IF NOT m_xInitial THEN
	BarCylinderIO.tLoadDelay:=T#3s;
	m_xInitial:=1;
END_IF;
IF g_xManual THEN    (*手动*)
	BarCylinderIO.xNextRun:=0;
	BarCylinderIO.xBarCylinder:=BarCylinderIO.xBarCylinderButton;
	BarCylinderIO.xBarCylinderSecondary	:=BarCylinderIO.xBarSecondaryButton;
	BarCylinderIO.xTransportMotorCW:= BarCylinderIO.xTransportMotorCWButton 
																	AND NOT BarCylinderIO.xTransportMotorCCWButton 
																	AND NOT BarCylinderIO.xTransportMotorCCW ;
	BarCylinderIO.xTransportMotorCCW:=BarCylinderIO.xTransportMotorCCWButton 
																		AND NOT BarCylinderIO.xTransportMotorCWButton 
																		AND NOT BarCylinderIO.xTransportMotorCW;
END_IF;
IF g_xAuto THEN(*自动*)
    IF BarCylinderIO.xUnload   (*下料*)
    	AND NOT BarCylinderIO.xEmpty  (*有料*)
    	AND NOT BarCylinderIO.xNextRun  (*下段线体旋转*)
    	AND NOT (g_xResetSingle AND BarCylinderIO.iDeviceID=g_iDeviceIDSelect)(*无复位信号*)
    	THEN(*收到卸料命令，当阻挡器不为空时*)
    	BarCylinderIO.xBarCylinder:=1;
    	BarCylinderIO.xNextRun:=1;(*确保下料命令只执行一次，防止物料在输送过程中又有卸料命令导致多次卸料*)
    	BarCylinderIO.xTransportMotorCW:=1;
    END_IF;
    IF NOT  BarCylinderIO.xUnload  THEN
    	BarCylinderIO.xNextRun:=0;
    	BarCylinderIO.xBarCylinder:=0;
    END_IF;
    m_tonLoadDelay(IN:= BarCylinderIO.xPresentSwitch ,PT:= BarCylinderIO.tLoadDelay ,Q:= m_xLoadDelay,ET:= m_tLoadDelayCurrentTime );
    IF m_xLoadDelay OR  BarCylinderIO.xNextRun  THEN
    	BarCylinderIO.xEmpty:=0;
    	BarCylinderIO.xBarCylinderSecondary:=1;
    ELSE
    	BarCylinderIO.xEmpty:=1;
    	BarCylinderIO.xBarCylinderSecondary:=0;
    END_IF;
    (*如果为空，气缸顶起*)
   IF  BarCylinderIO.xEmpty  THEN
   	   BarCylinderIO.xBarCylinder:=0;
   END_IF;
   	IF BarCylinderIO.xLoad AND BarCylinderIO.xEmpty  THEN
		BarCylinderIO.xTransportMotorCW:=1;
   	END_IF;  
   	IF (BarCylinderIO.xLoad=0 OR BarCylinderIO.xEmpty=0)  AND (BarCylinderIO.xUnload=0 OR BarCylinderIO.xEmpty) THEN
   		BarCylinderIO.xTransportMotorCW:=0;
   	END_IF;
END_IF;  
IF BarCylinderIO.xEmpty AND BarCylinderIO.xLoad=0 THEN
	BarCylinderIO.iProductCategory:=0;
END_IF;

IF NOT g_xEStop THEN
	 BarCylinderIO.xTransportMotorCW:=0;
	 BarCylinderIO.xTransportMotorCCW:=0;
	 BarCylinderIO.xBarCylinder:=0;
END_IF;

(*//复位*)
IF  (g_xResetSingle AND BarCylinderIO.iDeviceID=g_iDeviceIDSelect)THEN   (* //非正常情况下切断xNextRun不会复位，通过这个标志位会出发报警*)(*增加单体复位*)
	 BarCylinderIO.xNextRun:=0; 
END_IF;
END_FUNCTION_BLOCK
